// TIA Portal project "Bandsteuerung" (V20)

(* hardware
DEVICE "S7-1500/ET200MP station_1"  S7-1500 station
   slot 0: "Rail_0"  Rack  6ES7 590-1***0-0AA0
   slot 1: "PLC_2"  CPU 1511-1 PN  6ES7 511-1AK00-0AB0  V1.8
      slot 3: "CPU display_1"  6ES7591-1AA00-0AA0
      slot 32768: "PROFINET interface_1"  X1
         slot 32769: "Port_1"  X1 P1
         slot 32770: "Port_2"  X1 P2
*)

// ===== PLC "PLC_2"  CPU 1511-1 PN =====

VAR_GLOBAL   // PLC tag table "Default tag table"
   "S1" AT %I0.0 : Bool;   // START-TASTE BAND 1
   "S2" AT %I0.1 : Bool;   // START-TASTE BAND 2
   "S3" AT %I0.2 : Bool;   // STOP-TASTE BAND 1
   "S4" AT %I0.3 : Bool;   // STOP-TASTE BAND 2
   "M1" AT %Q0.0 : Bool;
   "M2" AT %Q0.1 : Bool;
   "M3" AT %Q0.2 : Bool;
   "Tag_1" AT %T1 : Timer;
   "Tag_2" AT %T2 : Timer;
   "Tag_3" AT %T3 : Timer;
   "M_Band1" AT %Q0.3 : Bool;
   "M_Band2" AT %Q0.4 : Bool;
END_VAR

// folder: System blocks/Program resources

DATA_BLOCK "IEC_Timer_0_DB"   // DB1
{ S7_Optimized_Access := 'TRUE' }
AUTHOR : Simatic
FAMILY : IEC
NAME : IEC_TMR
VERSION : 1.0
// stored: InstanceOfName IEC_TIMER
"IEC_TIMER"
BEGIN
END_DATA_BLOCK

DATA_BLOCK "IEC_Timer_0_DB_1"   // DB2
{ S7_Optimized_Access := 'TRUE' }
AUTHOR : Simatic
FAMILY : IEC
NAME : IEC_TMR
VERSION : 1.0
// stored: InstanceOfName IEC_TIMER
"IEC_TIMER"
BEGIN
END_DATA_BLOCK

DATA_BLOCK "IEC_Timer_0_DB_2"   // DB3
{ S7_Optimized_Access := 'TRUE' }
AUTHOR : Simatic
FAMILY : IEC
NAME : IEC_TMR
VERSION : 1.0
// stored: InstanceOfName IEC_TIMER
"IEC_TIMER"
BEGIN
END_DATA_BLOCK

// folder: (top level)

FUNCTION "FC_Bandsteuerung" : Void   // FC1, FBD
{ S7_Optimized_Access := 'FALSE' }
VERSION : 0.1
BEGIN

REGION Network 1: Turn ON Förderband 1 with condition of M2 being OFF
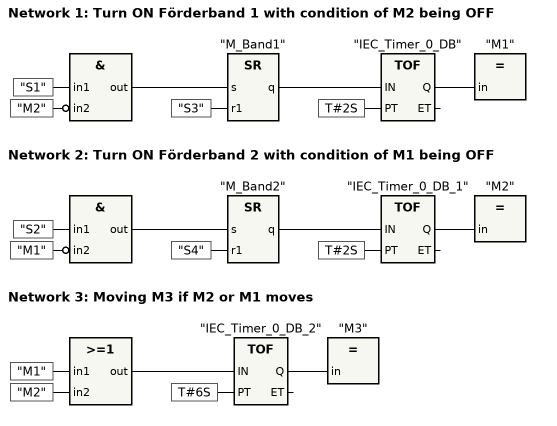
   IF "S1" AND NOT "M2" THEN
       "M_Band1" := TRUE;   // SR flip-flop
   END_IF;
   IF "S3" THEN "M_Band1" := FALSE; END_IF;
   "IEC_Timer_0_DB".TOF(IN := "M_Band1", PT := T#2S);
   "M1" := "IEC_Timer_0_DB".Q;
END_REGION

REGION Network 2: Turn ON Förderband 2 with condition of M1 being OFF
   IF "S2" AND NOT "M1" THEN
       "M_Band2" := TRUE;   // SR flip-flop
   END_IF;
   IF "S4" THEN "M_Band2" := FALSE; END_IF;
   "IEC_Timer_0_DB_1".TOF(IN := "M_Band2", PT := T#2S);
   "M2" := "IEC_Timer_0_DB_1".Q;
END_REGION

REGION Network 3: Moving M3 if M2 or M1 moves
   "IEC_Timer_0_DB_2".TOF(IN := "M1" OR "M2", PT := T#6S);
   "M3" := "IEC_Timer_0_DB_2".Q;
END_REGION
END_FUNCTION

ORGANIZATION_BLOCK "Main"   // OB1, LAD, ProgramCycle
TITLE = "Main Program Sweep (Cycle)"
{ S7_Optimized_Access := 'FALSE' }
VERSION : 0.1
   VAR_TEMP
      OB1_EV_CLASS : Byte;   // Bits 0-3 = 1 (Coming event), Bits 4-7 = 1 (Event class 1)
      OB1_SCAN_1 : Byte;   // 1 (Cold restart scan 1 of OB 1), 3 (Scan 2-n of OB 1)
      OB1_PRIORITY : Byte;   // Priority of OB Execution
      OB1_OB_NUMBR : Byte;   // 1 (Organization block 1, OB1)
      OB1_RESERVED_1 : Byte;   // Reserved for system
      OB1_RESERVED_2 : Byte;   // Reserved for system
      OB1_PREV_CYCLE : Int;   // Cycle time of previous OB1 scan (milliseconds)
      OB1_MIN_CYCLE : Int;   // Minimum cycle time of OB1 (milliseconds)
      OB1_MAX_CYCLE : Int;   // Maximum cycle time of OB1 (milliseconds)
      OB1_DATE_TIME : Date_And_Time;   // Date and time OB1 started
   END_VAR
BEGIN

REGION Network 1
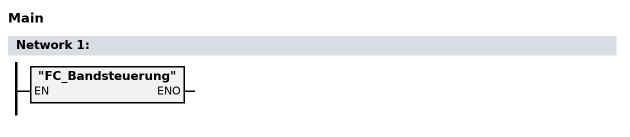
   RUNG wire#powerrail
      "FC_Bandsteuerung"()
   END_RUNG
   // the same network as SCL:
   "FC_Bandsteuerung"();
END_REGION
END_ORGANIZATION_BLOCK